// TIA Portal project "ProjectTest" (V15.1) (continued)
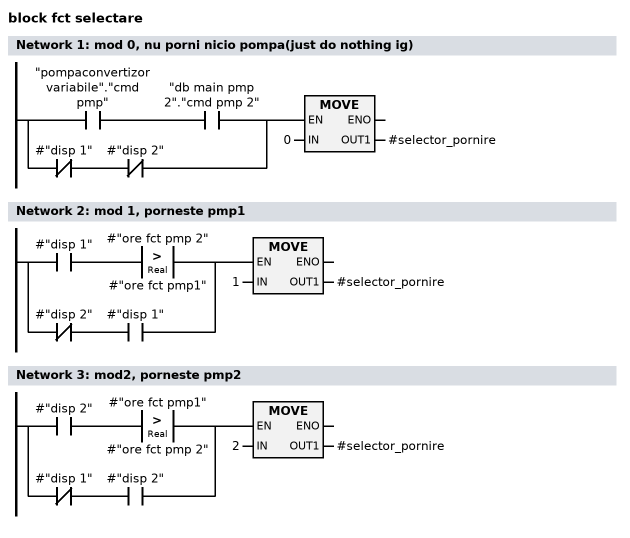
   RUNG wire#powerrail
      Contact( "pompaconvertizor variabile"."cmd pmp" )
      Contact( "db main pmp 2"."cmd pmp 2" )
      wire#w1
      Move(in := 0, out1 => #selector_pornire)
   END_RUNG
   RUNG wire#powerrail
      I_Contact( #"disp 1" )
      I_Contact( #"disp 2" )
   END_RUNG wire#w1
   // the same network as SCL:
   IF ("pompaconvertizor variabile"."cmd pmp" AND "db main pmp 2"."cmd pmp 2") OR (NOT #"disp 1" AND NOT #"disp 2") THEN
       #selector_pornire := 0;
   END_IF;
END_REGION

REGION Network 2: mod 1, porneste pmp1
   RUNG wire#powerrail
      Contact( #"disp 1" )
      { S7_Templates := "SrcType := Real" } GT_Contact(in1 := #"ore fct pmp 2", in2 := #"ore fct pmp1")
      wire#w1
      Move(in := 1, out1 => #selector_pornire)
   END_RUNG
   RUNG wire#powerrail
      I_Contact( #"disp 2" )
      Contact( #"disp 1" )
   END_RUNG wire#w1
   // the same network as SCL:
   IF (#"disp 1" AND (#"ore fct pmp 2" > #"ore fct pmp1")) OR (NOT #"disp 2" AND #"disp 1") THEN
       #selector_pornire := 1;
   END_IF;
END_REGION

REGION Network 3: mod2, porneste pmp2
   RUNG wire#powerrail
      Contact( #"disp 2" )
      { S7_Templates := "SrcType := Real" } GT_Contact(in1 := #"ore fct pmp1", in2 := #"ore fct pmp 2")
      wire#w1
      Move(in := 2, out1 => #selector_pornire)
   END_RUNG
   RUNG wire#powerrail
      I_Contact( #"disp 1" )
      Contact( #"disp 2" )
   END_RUNG wire#w1
   // the same network as SCL:
   IF (#"disp 2" AND (#"ore fct pmp1" > #"ore fct pmp 2")) OR (NOT #"disp 1" AND #"disp 2") THEN
       #selector_pornire := 2;
   END_IF;
END_REGION
END_FUNCTION_BLOCK

FUNCTION_BLOCK "pompa convertizor"   // FB2, LAD
{ S7_Optimized_Access := 'TRUE' }
VERSION : 0.1
   VAR_INPUT
      int_pid : Real;
      disponibil : Bool;
      mad_fct : Bool;
      fault : Bool;
      ESD : Bool;
      B_start_manual : Bool;
      B_stop_manual : Bool;
      viteza_impusa_manual : Real;
      start_auto : Bool;
   END_VAR
   VAR_OUTPUT
      out_debit : Real;
      cmd_pompa : Bool;
   END_VAR
   VAR
      reg_auto : Bool;
      reg_man : Bool;
   END_VAR
BEGIN

REGION Network 1: selctare regim auto
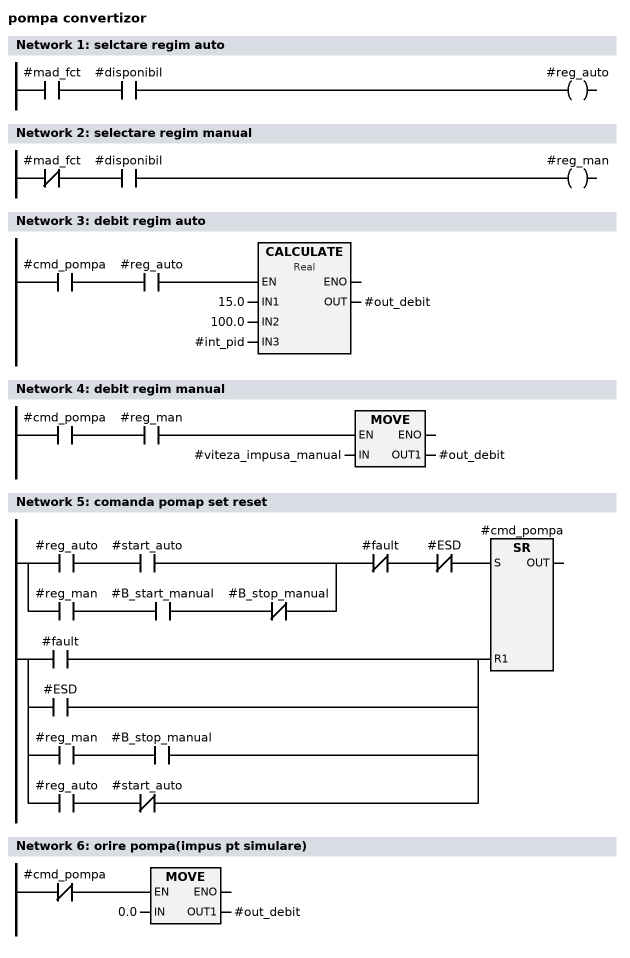
   RUNG wire#powerrail
      Contact( #mad_fct )
      Contact( #disponibil )
      Coil( #reg_auto )
   END_RUNG
   // the same network as SCL:
   #reg_auto := #mad_fct AND #disponibil;
END_REGION

REGION Network 2: selectare regim manual
   RUNG wire#powerrail
      I_Contact( #mad_fct )
      Contact( #disponibil )
      Coil( #reg_man )
   END_RUNG
   // the same network as SCL:
   #reg_man := NOT #mad_fct AND #disponibil;
END_REGION

REGION Network 3: debit regim auto
   RUNG wire#powerrail
      Contact( #cmd_pompa )
      Contact( #reg_auto )
      { S7_Templates := "SrcType := Real"; S7_Expression := "IN1 * IN3 / IN2" } Calculate(in1 := 15.0, in2 := 100.0, in3 := #int_pid, out => #out_debit)
   END_RUNG
   // the same network as SCL:
   IF #cmd_pompa AND #reg_auto THEN #out_debit := 15.0 * #int_pid / 100.0; END_IF;
END_REGION

REGION Network 4: debit regim manual
   RUNG wire#powerrail
      Contact( #cmd_pompa )
      Contact( #reg_man )
      Move(in := #viteza_impusa_manual, out1 => #out_debit)
   END_RUNG
   // the same network as SCL:
   IF #cmd_pompa AND #reg_man THEN #out_debit := #viteza_impusa_manual; END_IF;
END_REGION

REGION Network 5: comanda pomap set reset
   RUNG wire#powerrail
      Contact( #reg_auto )
      Contact( #start_auto )
      wire#w1
      I_Contact( #fault )
      I_Contact( #ESD )
      S_SR(operand := #cmd_pompa, r1 := wire#w2)
   END_RUNG
   RUNG wire#powerrail
      Contact( #reg_man )
      Contact( #B_start_manual )
      I_Contact( #B_stop_manual )
   END_RUNG wire#w1
   RUNG wire#powerrail
      Contact( #fault )
   END_RUNG wire#w2
   RUNG wire#powerrail
      Contact( #ESD )
   END_RUNG wire#w2
   RUNG wire#powerrail
      Contact( #reg_man )
      Contact( #B_stop_manual )
   END_RUNG wire#w2
   RUNG wire#powerrail
      Contact( #reg_auto )
      I_Contact( #start_auto )
   END_RUNG wire#w2
   // the same network as SCL:
   IF ((#reg_auto AND #start_auto) OR (#reg_man AND #B_start_manual AND NOT #B_stop_manual)) AND NOT #fault AND NOT #ESD THEN
       #cmd_pompa := TRUE;   // SR flip-flop
   END_IF;
   IF #fault OR #ESD OR (#reg_man AND #B_stop_manual) OR (#reg_auto AND NOT #start_auto) THEN
       #cmd_pompa := FALSE;
   END_IF;
END_REGION

REGION Network 6: orire pompa(impus pt simulare)
   RUNG wire#powerrail
      I_Contact( #cmd_pompa )
      Move(in := 0.0, out1 => #out_debit)
   END_RUNG
   // the same network as SCL:
   IF NOT #cmd_pompa THEN #out_debit := 0.0; END_IF;
END_REGION
END_FUNCTION_BLOCK

ORGANIZATION_BLOCK "Main"   // OB1, LAD, ProgramCycle
TITLE = "Main Program Sweep (Cycle)"
{ S7_Optimized_Access := 'TRUE' }
VERSION : 0.1
   VAR_INPUT
      Initial_Call : Bool;   // Initial call of this OB
      Remanence : Bool;   // =True, if remanent data are available
   END_VAR
   VAR_TEMP   // added for the SCL form of the ladder/FBD networks
      _w1 : Bool;
      _w2 : Bool;
      _w3 : Bool;
      _w4 : Bool;
   END_VAR
BEGIN

REGION Network 1: initializare pompe cu convertizoare
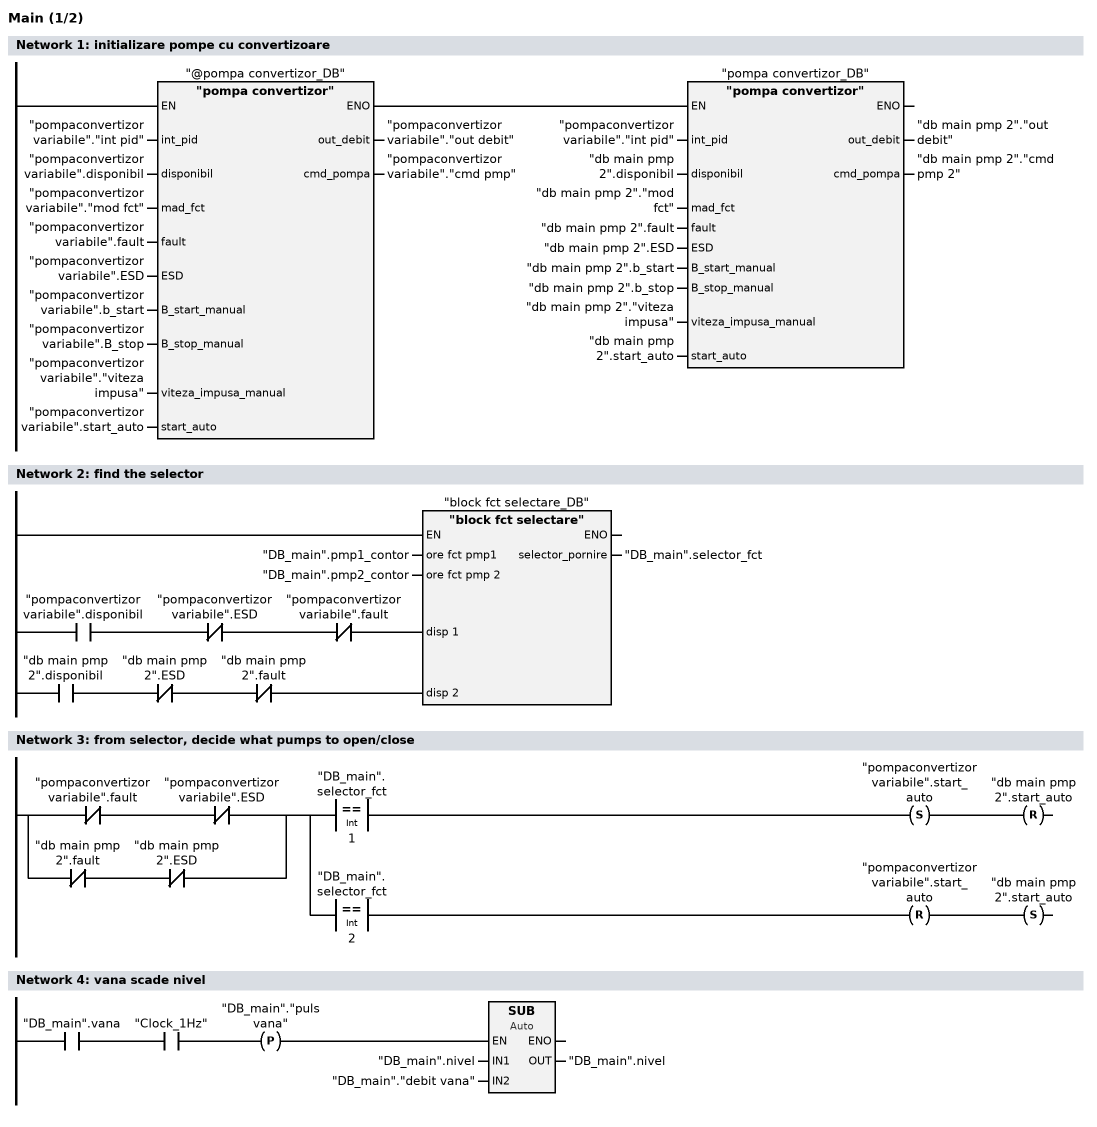
   RUNG wire#powerrail
      "@pompa convertizor_DB"(int_pid := "pompaconvertizor variabile"."int pid", disponibil := "pompaconvertizor variabile".disponibil, mad_fct := "pompaconvertizor variabile"."mod fct", fault := "pompaconvertizor variabile".fault, ESD := "pompaconvertizor variabile".ESD, B_start_manual := "pompaconvertizor variabile".b_start, B_stop_manual := "pompaconvertizor variabile".B_stop, viteza_impusa_manual := "pompaconvertizor variabile"."viteza impusa", start_auto := "pompaconvertizor variabile".start_auto, out_debit => "pompaconvertizor variabile"."out debit", cmd_pompa => "pompaconvertizor variabile"."cmd pmp")
      "pompa convertizor_DB"(int_pid := "pompaconvertizor variabile"."int pid", disponibil := "db main pmp 2".disponibil, mad_fct := "db main pmp 2"."mod  fct", fault := "db main pmp 2".fault, ESD := "db main pmp 2".ESD, B_start_manual := "db main pmp 2".b_start, B_stop_manual := "db main pmp 2".b_stop, viteza_impusa_manual := "db main pmp 2"."viteza impusa", start_auto := "db main pmp 2".start_auto, out_debit => "db main pmp 2"."out debit", cmd_pompa => "db main pmp 2"."cmd pmp 2")
   END_RUNG
   // the same network as SCL:
   "@pompa convertizor_DB"(int_pid := "pompaconvertizor variabile"."int pid",   // "pompa convertizor"
                           disponibil := "pompaconvertizor variabile".disponibil,
                           mad_fct := "pompaconvertizor variabile"."mod fct",
                           fault := "pompaconvertizor variabile".fault,
                           ESD := "pompaconvertizor variabile".ESD,
                           B_start_manual := "pompaconvertizor variabile".b_start,
                           B_stop_manual := "pompaconvertizor variabile".B_stop,
                           viteza_impusa_manual := "pompaconvertizor variabile"."viteza impusa",
                           start_auto := "pompaconvertizor variabile".start_auto,
                           out_debit => "pompaconvertizor variabile"."out debit",
                           cmd_pompa => "pompaconvertizor variabile"."cmd pmp",
                           ENO => #_w1);
   IF #_w1 THEN
       "pompa convertizor_DB"(int_pid := "pompaconvertizor variabile"."int pid",   // "pompa convertizor"
                              disponibil := "db main pmp 2".disponibil,
                              mad_fct := "db main pmp 2"."mod  fct",
                              fault := "db main pmp 2".fault,
                              ESD := "db main pmp 2".ESD,
                              B_start_manual := "db main pmp 2".b_start,
                              B_stop_manual := "db main pmp 2".b_stop,
                              viteza_impusa_manual := "db main pmp 2"."viteza impusa",
                              start_auto := "db main pmp 2".start_auto,
                              out_debit => "db main pmp 2"."out debit",
                              cmd_pompa => "db main pmp 2"."cmd pmp 2");
   END_IF;
END_REGION

REGION Network 2: find the selector
   RUNG wire#powerrail
      "block fct selectare_DB"("disp 1" := wire#w1, "disp 2" := wire#w2, "ore fct pmp1" := "DB_main".pmp1_contor, "ore fct pmp 2" := "DB_main".pmp2_contor, selector_pornire => "DB_main".selector_fct)
   END_RUNG
   RUNG wire#powerrail
      Contact( "pompaconvertizor variabile".disponibil )
      I_Contact( "pompaconvertizor variabile".ESD )
      I_Contact( "pompaconvertizor variabile".fault )
   END_RUNG wire#w1
   RUNG wire#powerrail
      Contact( "db main pmp 2".disponibil )
      I_Contact( "db main pmp 2".ESD )
      I_Contact( "db main pmp 2".fault )
   END_RUNG wire#w2
   // the same network as SCL:
   "block fct selectare_DB"("ore fct pmp1" := "DB_main".pmp1_contor,   // "block fct selectare"
                           "ore fct pmp 2" := "DB_main".pmp2_contor,
                           "disp 1" := "pompaconvertizor variabile".disponibil AND NOT "pompaconvertizor variabile".ESD AND NOT "pompaconvertizor variabile".fault,
                           "disp 2" := "db main pmp 2".disponibil AND NOT "db main pmp 2".ESD AND NOT "db main pmp 2".fault,
                           selector_pornire => "DB_main".selector_fct);
END_REGION

REGION Network 3: from selector, decide what pumps to open/close
   RUNG wire#powerrail
      I_Contact( "pompaconvertizor variabile".fault )
      I_Contact( "pompaconvertizor variabile".ESD )
      wire#w1
      { S7_Templates := "SrcType := Int" } EQ_Contact(in1 := "DB_main".selector_fct, in2 := 1)
      S_Coil( "pompaconvertizor variabile".start_auto )
      R_Coil( "db main pmp 2".start_auto )
   END_RUNG
   RUNG wire#powerrail
      I_Contact( "db main pmp 2".fault )
      I_Contact( "db main pmp 2".ESD )
   END_RUNG wire#w1
   RUNG wire#w1
      { S7_Templates := "SrcType := Int" } EQ_Contact(in1 := "DB_main".selector_fct, in2 := 2)
      R_Coil( "pompaconvertizor variabile".start_auto )
      S_Coil( "db main pmp 2".start_auto )
   END_RUNG
   // the same network as SCL:
   #_w1 := (NOT "pompaconvertizor variabile".fault AND NOT "pompaconvertizor variabile".ESD) OR (NOT "db main pmp 2".fault AND NOT "db main pmp 2".ESD);
   IF #_w1 AND ("DB_main".selector_fct = 1) THEN
       "pompaconvertizor variabile".start_auto := TRUE;
       "db main pmp 2".start_auto := FALSE;
   END_IF;
   IF #_w1 AND ("DB_main".selector_fct = 2) THEN
       "pompaconvertizor variabile".start_auto := FALSE;
       "db main pmp 2".start_auto := TRUE;
   END_IF;
END_REGION

REGION Network 4: vana scade nivel
   RUNG wire#powerrail
      Contact( "DB_main".vana )
      Contact( "Clock_1Hz" )
      P_Trig( "DB_main"."puls vana" )
      Sub(in1 := "DB_main".nivel, in2 := "DB_main"."debit vana", out => "DB_main".nivel)
   END_RUNG
   // the same network as SCL:
   #_w1 := "DB_main".vana AND "Clock_1Hz";
   #_w2 := #_w1 AND NOT "DB_main"."puls vana";   // rising edge
   "DB_main"."puls vana" := #_w1;
   IF #_w2 THEN "DB_main".nivel := "DB_main".nivel - "DB_main"."debit vana"; END_IF;
END_REGION

REGION Network 5: pompe add la nivel
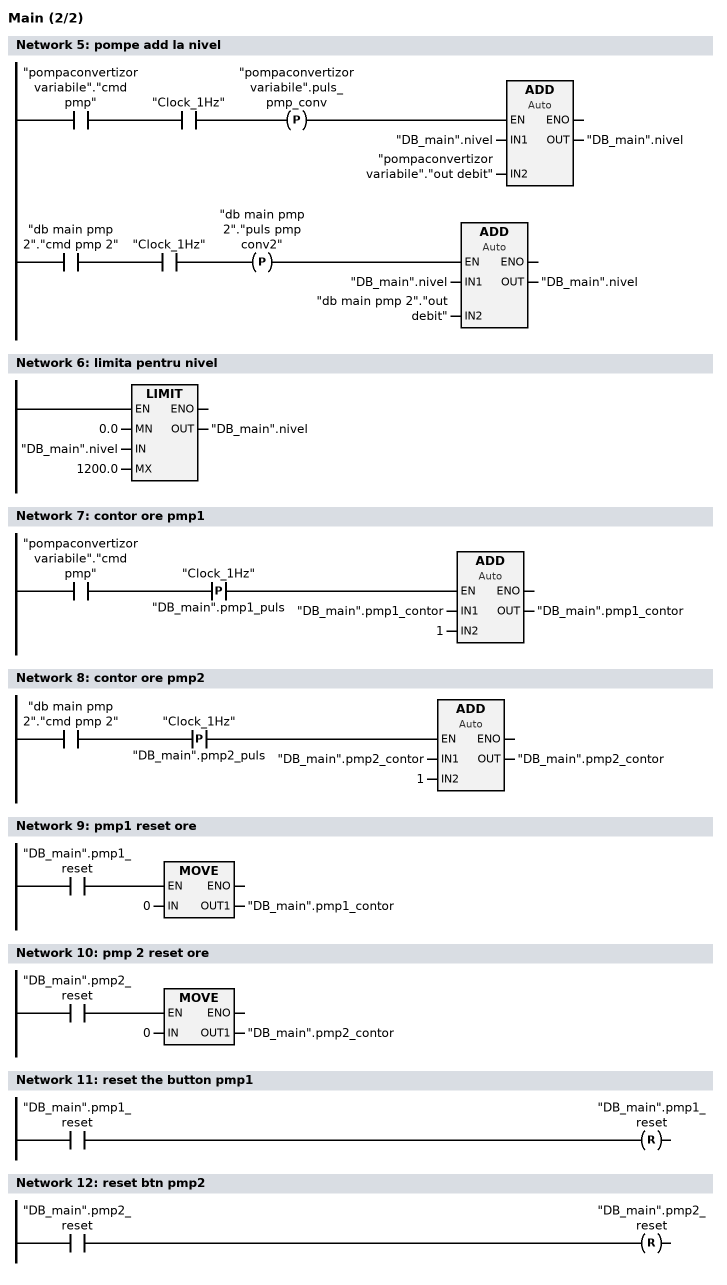
   RUNG wire#powerrail
      Contact( "pompaconvertizor variabile"."cmd pmp" )
      Contact( "Clock_1Hz" )
      P_Trig( "pompaconvertizor variabile".puls_pmp_conv )
      Add(in1 := "DB_main".nivel, in2 := "pompaconvertizor variabile"."out debit", out => "DB_main".nivel)
   END_RUNG
   RUNG wire#powerrail
      Contact( "db main pmp 2"."cmd pmp 2" )
      Contact( "Clock_1Hz" )
      P_Trig( "db main pmp 2"."puls pmp conv2" )
      Add(in1 := "DB_main".nivel, in2 := "db main pmp 2"."out debit", out => "DB_main".nivel)
   END_RUNG
   // the same network as SCL:
   #_w1 := "pompaconvertizor variabile"."cmd pmp" AND "Clock_1Hz";
   #_w2 := #_w1 AND NOT "pompaconvertizor variabile".puls_pmp_conv;   // rising edge
   "pompaconvertizor variabile".puls_pmp_conv := #_w1;
   IF #_w2 THEN "DB_main".nivel := "DB_main".nivel + "pompaconvertizor variabile"."out debit"; END_IF;
   #_w3 := "db main pmp 2"."cmd pmp 2" AND "Clock_1Hz";
   #_w4 := #_w3 AND NOT "db main pmp 2"."puls pmp conv2";   // rising edge
   "db main pmp 2"."puls pmp conv2" := #_w3;
   IF #_w4 THEN "DB_main".nivel := "DB_main".nivel + "db main pmp 2"."out debit"; END_IF;
END_REGION

REGION Network 6: limita pentru nivel
   "DB_main".nivel := LIMIT(MN := 0.0, IN := "DB_main".nivel, MX := 1200.0);
END_REGION

REGION Network 7: contor ore pmp1
   RUNG wire#powerrail
      Contact( "pompaconvertizor variabile"."cmd pmp" )
      P_Contact(operand := "Clock_1Hz", bit := "DB_main".pmp1_puls)
      Add(in1 := "DB_main".pmp1_contor, in2 := 1, out => "DB_main".pmp1_contor)
   END_RUNG
   // the same network as SCL:
   #_w1 := "pompaconvertizor variabile"."cmd pmp" AND "Clock_1Hz" AND NOT "DB_main".pmp1_puls;   // rising edge of "Clock_1Hz"
   "DB_main".pmp1_puls := "Clock_1Hz";
   IF #_w1 THEN "DB_main".pmp1_contor := "DB_main".pmp1_contor + 1; END_IF;
END_REGION

REGION Network 8: contor ore pmp2
   RUNG wire#powerrail
      Contact( "db main pmp 2"."cmd pmp 2" )
      P_Contact(operand := "Clock_1Hz", bit := "DB_main".pmp2_puls)
      Add(in1 := "DB_main".pmp2_contor, in2 := 1, out => "DB_main".pmp2_contor)
   END_RUNG
   // the same network as SCL:
   #_w1 := "db main pmp 2"."cmd pmp 2" AND "Clock_1Hz" AND NOT "DB_main".pmp2_puls;   // rising edge of "Clock_1Hz"
   "DB_main".pmp2_puls := "Clock_1Hz";
   IF #_w1 THEN "DB_main".pmp2_contor := "DB_main".pmp2_contor + 1; END_IF;
END_REGION

REGION Network 9: pmp1 reset ore
   RUNG wire#powerrail
      Contact( "DB_main".pmp1_reset )
      Move(in := 0, out1 => "DB_main".pmp1_contor)
   END_RUNG
   // the same network as SCL:
   IF "DB_main".pmp1_reset THEN "DB_main".pmp1_contor := 0; END_IF;
END_REGION

REGION Network 10: pmp 2 reset ore
   RUNG wire#powerrail
      Contact( "DB_main".pmp2_reset )
      Move(in := 0, out1 => "DB_main".pmp2_contor)
   END_RUNG
   // the same network as SCL:
   IF "DB_main".pmp2_reset THEN "DB_main".pmp2_contor := 0; END_IF;
END_REGION

REGION Network 11: reset the button pmp1
   RUNG wire#powerrail
      Contact( "DB_main".pmp1_reset )
      R_Coil( "DB_main".pmp1_reset )
   END_RUNG
   // the same network as SCL:
   IF "DB_main".pmp1_reset THEN "DB_main".pmp1_reset := FALSE; END_IF;
END_REGION

REGION Network 12: reset btn pmp2
   RUNG wire#powerrail
      Contact( "DB_main".pmp2_reset )
      R_Coil( "DB_main".pmp2_reset )
   END_RUNG
   // the same network as SCL:
   IF "DB_main".pmp2_reset THEN "DB_main".pmp2_reset := FALSE; END_IF;
END_REGION
END_ORGANIZATION_BLOCK

ORGANIZATION_BLOCK "Cyclic for pid"   // OB30, LAD, CyclicInterrupt
{ S7_Optimized_Access := 'TRUE' }
VERSION : 0.1
   VAR_INPUT
      Initial_Call : Bool;   // Initial call of this OB
      Event_Count : Int;   // Events discarded
   END_VAR
BEGIN

REGION Network 1
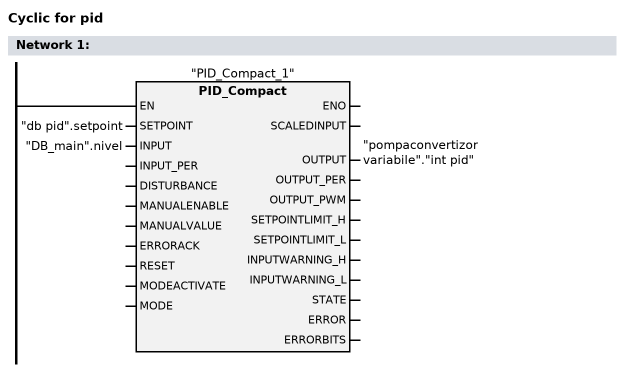
   "PID_Compact_1"(Setpoint := "db pid".setpoint,   // PID_Compact
                   Input := "DB_main".nivel,
                   Output => "pompaconvertizor variabile"."int pid");
END_REGION
END_ORGANIZATION_BLOCK

(* ===== HMI "HMI_RT_1" =====
system functions are stored by id; their names below are inferred from use
connection "HMI_Connection_1": ETHERNET, SMART_S7_1200_OMS

HMI tags "Default tag table"
   "Bazin_Nivel" : Real = PLC Bazin.Nivel, 1 s
   "Bazin_Vana golire" : Bool = PLC Bazin."Vana golire", 1 s
   "Pompa_1_Contor" : UInt = PLC Pompa_1.Contor, 1 s
   "Pompa_2_Contor" : UInt = PLC Pompa_2.Contor, 1 s
   "Pompa_1_Reset" : Bool = PLC Pompa_1.Reset, 1 s
   "Pompa_2_Reset" : Bool = PLC Pompa_2.Reset, 1 s
   "Bazin_Cheie" : Int = PLC Bazin.Cheie, 1 s
   "Pompa1" : Bool = PLC Pompa1 AT %Q0.0, 1 s
   "Pompa2" : Bool = PLC Pompa2 AT %Q0.1, 1 s

screen "Screen_1" 800x480
   Bar "Bar_1" at 259,52 size 164x377; MinimumValue 0; MaximumValue 1000
      ProcessValue <- "Bazin_Nivel"
   Button "Button_1" at 85,411 size 96x32; TextOff 'Reset vana'
      on Click: SetBit("Bazin_Vana golire")
   IOField "I/O field_1" at 480,77 size 96x32; FormatPattern 99999; Unit s
      ProcessValue <- "Pompa_1_Contor"
   TextField "Text field_1" at 480,53 size 96x20; Text 'Counter pmp1'
   IOField "I/O field_2" at 486,154 size 96x32; FormatPattern 99999; Unit s
      ProcessValue <- "Pompa_2_Contor"
   TextField "Text field_2" at 486,134 size 96x20; Text 'Counter pmp2'
   Button "Button_2" at 610,78 size 96x32; TextOff 'Reset1'
      on Click: SetBit("Pompa_1_Reset")
   Button "Button_3" at 609,153 size 96x32; TextOff 'Reset2'
      on Activate: SetBit("Pompa_2_Reset")
   Button "Button_4" at 56,117 size 96x32; TextOff '0'
      on Click: SetTag("Bazin_Cheie", 0)
   Button "Button_5" at 56,185 size 96x32; TextOff '1'
      on Click: SetTag("Bazin_Cheie", 1)
   Button "Button_6" at 56,250 size 96x32; TextOff '2'
      on Click: SetTag("Bazin_Cheie", 2)
   TextField "Text field_3" at 65,67 size 70x20; Text 'Set config'
   Rectangle "Rectangle_1" at 85,351 size 96x48
      Appearance <- "Bazin_Vana golire"
   Circle "Circle_1" at 505,319 size 48x48
      Appearance <- "Pompa1"
   Circle "Circle_2" at 593,321 size 48x48
      Appearance <- "Pompa2"
   TextField "Text field_4" at 505,299 size 40x20; Text 'Pmp1'
   TextField "Text field_5" at 593,302 size 40x20; Text 'Pmp2'
   Button "Button_7" at 610,223 size 96x32; TextOff 'doar reset'
*)

(* ===== HMI "HMI_RT_2" =====
system functions are stored by id; their names below are inferred from use
connection "HMI_Connection_2": ETHERNET, SMART_S7_1500_OMS

HMI tags "Default tag table"
   "Tag_ScreenNumber" : UInt, internal
   "DB_main_nivel" : Real = PLC DB_main.nivel, 1 s
   "DB_main_pmp1_contor" : Int = PLC DB_main.pmp1_contor, 1 s
   "DB_main_pmp2_contor" : Int = PLC DB_main.pmp2_contor, 1 s
   "pompaconvertizor variabile_int pid" : Real = PLC "pompaconvertizor variabile"."int pid", 1 s
   "DB_main_selector_fct" : Int = PLC DB_main.selector_fct, 1 s
   "db pid_setpoint" : Real = PLC "db pid".setpoint, 1 s
   "DB_main_pmp1_reset" : Bool = PLC DB_main.pmp1_reset, 1 s
   "DB_main_pmp2_reset" : Bool = PLC DB_main.pmp2_reset, 1 s
   "DB_main_vana" : Bool = PLC DB_main.vana, 1 s
   "pompaconvertizor variabile_fault" : Bool = PLC "pompaconvertizor variabile".fault, 1 s
   "pompaconvertizor variabile_ESD" : Bool = PLC "pompaconvertizor variabile".ESD, 1 s
   "db main pmp 2_fault" : Bool = PLC "db main pmp 2".fault, 1 s
   "db main pmp 2_ESD" : Bool = PLC "db main pmp 2".ESD, 1 s
   "pompaconvertizor variabile_start_auto" : Bool = PLC "pompaconvertizor variabile".start_auto, 1 s
   "db main pmp 2_start_auto" : Bool = PLC "db main pmp 2".start_auto, 1 s
   "pompaconvertizor variabile_out debit" : Real = PLC "pompaconvertizor variabile"."out debit", 1 s
   "db main pmp 2_out debit" : Real = PLC "db main pmp 2"."out debit", 1 s

Template "Template_1" 800x480
   Button "Exit" at 722,440 size 55x39; TextOff 'Exit'; PictureOff "ExitRuntime_KTP900_Basic_PN_TR"; PictureOn "ExitRuntime_KTP900_Basic_PN_TR"
      on Release: StopRuntime(0)
   Button "Template_Button" at 622,440 size 55x39; TextOff 'Text'
   Button "Template_Button_1" at 522,440 size 55x39; TextOff 'Text'
   Button "Template_Button_2" at 422,440 size 55x39; TextOff 'Text'
   Button "Template_Button_3" at 322,440 size 55x39; TextOff 'Text'
   Button "Template_Button_4" at 222,440 size 55x39; TextOff 'Text'
   Button "Alarms" at 122,440 size 55x39; TextOff 'Alarms'; PictureOff "AlarmDisplay_KTP900_Basic_PN_TR"; PictureOn "AlarmDisplay_KTP900_Basic_PN_TR"
      on Release: function_ef3f5d25("Alarm window_Unacknowledged", -1)
   Button "Start screen" at 22,440 size 55x39; TextOff 'Start screen'; PictureOff "NavigateHome_KTP900_Basic_PN_TR"; PictureOn "NavigateHome_KTP900_Basic_PN_TR"
      on Release: ActivateScreen("Root screen", 0)
   SymbolicIOField "Symbolic_IO_Field_Screen" at 73,7 size 620x26; TextOff '0'; TextOn '1'; TextList "TextList_ScreenNames"
      ProcessValue <- "Tag_ScreenNumber"
      on Change: ActivateScreenByNumber("Tag_ScreenNumber", 0)
   DateTimeField "HmiScreenItemData" at 695,20 size 105x20
   DateTimeField "HmiScreenItemData_1" at 695,0 size 105x20
   GraphicView "Logo" at 0,0 size 71x40; Picture "Logo of HMI_2"

screen "Root screen" 800x480, template "Template_1"
   on GenerateScreen: SetTag("Tag_ScreenNumber", 1)
   Bar "Bar_1" at 19,69 size 100x367; MinimumValue 0; MaximumValue 1000
      ProcessValue <- "DB_main_nivel"
   IOField "I/O field_1" at 182,69 size 96x32; FormatPattern 99999; Unit s
      ProcessValue <- "DB_main_pmp1_contor"
   IOField "I/O field_2" at 182,114 size 96x32; FormatPattern 99999; Unit s
      ProcessValue <- "DB_main_pmp2_contor"
   TextField "Text field_1" at 153,69 size 21x20; Text 'C1'
   TextField "Text field_2" at 153,118 size 21x20; Text 'C2'
   Button "Button_1" at 297,70 size 58x32; TextOff 'Reset 1'
      on Click: SetBit("DB_main_pmp1_reset")
   Button "Button_2" at 298,114 size 58x32; TextOff 'Reset 2'
      on Click: SetBit("DB_main_pmp2_reset")
   IOField "I/O field_3" at 182,157 size 96x32; FormatPattern 999; Unit %
      ProcessValue <- "pompaconvertizor variabile_int pid"
   TextField "Text field_3" at 137,159 size 42x20; Text 'Pid %'
   Button "Button_3" at 298,159 size 76x32; TextOff 'Reset vana'
      on Click: SetBit("DB_main_vana")
   IOField "I/O field_4" at 183,208 size 96x32; FormatPattern 9
      ProcessValue <- "DB_main_selector_fct"
   TextField "Text field_4" at 143,211 size 32x20; Text 'Mod'
   IOField "I/O field_5" at 183,279 size 96x32; FormatPattern 9999
      ProcessValue <- "db pid_setpoint"
   TextField "Text field_5" at 182,261 size 86x20; Text 'Setpoint PID'
   Button "Button_4" at 567,65 size 64x32; TextOff 'fault 1'
      on Click: SetBit("pompaconvertizor variabile_fault")
   Button "Button_5" at 660,106 size 64x32; TextOff 'ESD 2'
      on Click: SetBit("db main pmp 2_ESD")
   Button "Button_6" at 567,107 size 64x32; TextOff 'ESD 1'
      on Click: SetBit("pompaconvertizor variabile_ESD")
   Button "Button_7" at 662,63 size 62x32; TextOff 'fault 2'
      on Click: SetBit("db main pmp 2_fault")
   Circle "Circle_1" at 510,51 size 39x39
      Appearance <- "pompaconvertizor variabile_fault"
   Circle "Circle_2" at 744,106 size 39x39
      Appearance <- "db main pmp 2_ESD"
   Circle "Circle_3" at 736,50 size 39x39
      Appearance <- "db main pmp 2_fault"
   Circle "Circle_4" at 510,100 size 39x39
      Appearance <- "pompaconvertizor variabile_ESD"
   Circle "Circle_5" at 298,221 size 58x58
      Appearance <- "pompaconvertizor variabile_start_auto"
   Circle "Circle_6" at 299,291 size 58x58
      Appearance <- "db main pmp 2_start_auto"
   TextField "Text field_6" at 300,202 size 21x20; Text 'P1'
   TextField "Text field_7" at 289,271 size 21x20; Text 'P2'
   Circle "Circle_7" at 382,150 size 39x39
      Appearance <- "DB_main_vana"
   Button "Button_8" at 169,403 size 50x32; TextOff 'Just is'
   IOField "I/O field_6" at 183,334 size 96x32; FormatPattern 9999.99
      ProcessValue <- "DB_main_nivel"
   TextField "Text field_8" at 135,335 size 35x20; Text 'Nivel'
   Button "Button_9" at 587,33 size 26x32; TextOff 'r f'
      on Click: ResetBit("pompaconvertizor variabile_fault")
   Button "Button_10" at 674,137 size 26x32; TextOff 'r f'
      on Click: ResetBit("db main pmp 2_ESD")
   Button "Button_11" at 587,137 size 26x32; TextOff 'r f'
      on Click: ResetBit("pompaconvertizor variabile_ESD")
   Button "Button_12" at 678,31 size 26x32; TextOff 'r f'
      on Click: ResetBit("db main pmp 2_fault")
   Button "Button_13" at 555,255 size 96x32; TextOff 'Screen PID'
      on Activate: ActivateScreen("Screen_1", 0)

screen "Screen_1" 800x480
   TrendView "Trend view_1" at 89,11 size 691x400
   Button "Button_1" at 24,434 size 96x32; TextOff 'Screen main'
      on Activate: ActivateScreen("Root screen", 0)
*)